VERSION : 0.1
   VAR_INPUT
      search_term : WString;
      search_array : Array[*] of WString[1];
   END_VAR
   VAR_TEMP
      _i : Int;
      _length_search_array : UDInt;
   END_VAR
BEGIN
   #_length_search_array := "Array.Any.Length"(#search_array);
   FOR #_i := 0 TO UDINT_TO_INT(#_length_search_array - 1) DO
       IF #search_term = #search_array[#_i] THEN
           #"Array.WString.Is_Element" := TRUE;
           RETURN;
       END_IF;
   END_FOR;
   #"Array.WString.Is_Element" := FALSE;
END_FUNCTION

FUNCTION "Array.Int.First_Occurance" : DInt   // FC220, SCL
{ S7_Optimized_Access := 'TRUE' }
VERSION : 0.1
   VAR_INPUT
      int_array : Array[*] of Int;
      search_term : Int;
   END_VAR
   VAR_TEMP
      _i : DInt;
      _length : UDInt;
   END_VAR
BEGIN
   REGION "NOTES"
       (* 
       This function returns the first occurance of the search term.
       This function meant for use with collapsed arrays.
       See "Array.Int.Collapse" for collapse functionality.
       *)
   END_REGION


   REGION "GET LENGTH OF INPUT ARRAY"
       #_length := "Array.Any.Length"(#int_array);
   END_REGION


   REGION "FIND FIRST SEARCH TERM, -1 IF NONE"
       (*
       Its worth noting that "Array.Int.Is_Element" could return the index of the search term
       as an output, saving the processor some work. 
       The rework is justified by increased encapsulation.
       The time complexity for "Array.Int.First_Occurance" remains O(n).
       *)
       IF NOT "Array.Int.Is_Element"(int_array := #int_array, search_term := #search_term) THEN
           #"Array.Int.First_Occurance" := -1;
           RETURN;
       END_IF;
       WHILE #int_array[#_i] <> #search_term AND DINT_TO_UDINT(#_i) < #_length DO
           #_i += 1;
       END_WHILE;
   END_REGION


   REGION _name_
       #"Array.Int.First_Occurance" := #_i;
   END_REGION
END_FUNCTION

FUNCTION "Array.WString.Fill" : Void   // FC243, SCL
{ S7_Optimized_Access := 'TRUE' }
VERSION : 0.1
   VAR_INPUT
      value : WString;
   END_VAR
   VAR_IN_OUT
      "array" : Array[*] of WString;
   END_VAR
   VAR_TEMP
      _length : Int;
      _i : Int;
   END_VAR
BEGIN
   #_length := UDINT_TO_INT("Array.Any.Length"(#array)) - 1;
   FOR #_i := 0 TO #_length DO
       #array[#_i] := #value;
   END_FOR;
   RETURN;
END_FUNCTION

FUNCTION "Array.WString.Search" : Int   // FC244, SCL
{ S7_Optimized_Access := 'TRUE' }
VERSION : 0.1
   VAR_INPUT
      "array" : Array[*] of WString;
      search_term : WString;
   END_VAR
   VAR_TEMP
      _i : Int;
      _length : Int;
   END_VAR
   // Ret_Val : index of search term. returns -1 if not found.
BEGIN
   REGION "SEARCH ARRAY"
       #_length := UDINT_TO_INT("Array.Any.Length"(#array)) - 1;
       FOR #_i := 0 TO #_length DO
           IF #array[#_i] <> #search_term THEN
               CONTINUE;
           END_IF;
           #"Array.WString.Search" := #_i;
           RETURN;
       END_FOR;
   END_REGION

   REGION "RETURN"
       #"Array.WString.Search" := "NULL_TOKEN";
       RETURN;
   END_REGION
END_FUNCTION

// folder: Utilities/Bool

FUNCTION "Bool.Animate" : USInt   // FC9, SCL
{ S7_Optimized_Access := 'TRUE' }
VERSION : 0.1
   VAR_INPUT
      true_color : USInt;
      false_color : USInt;
      evaluation_signal : Bool;
   END_VAR
   VAR_TEMP
      animate : USInt;
   END_VAR
BEGIN
   REGION "FALSE COLOR"
       IF NOT #evaluation_signal THEN
           #animate := #false_color;
       END_IF;
   END_REGION

   REGION "TRUE COLOR"
       IF #evaluation_signal THEN
           #animate := #true_color;
       END_IF;
   END_REGION

   REGION "FUNCTION RETURN"
       #"Bool.Animate" := #animate;
   END_REGION
END_FUNCTION

FUNCTION "Bool.Rising_Edge" : Bool   // FC177, SCL
{ S7_Optimized_Access := 'TRUE' }
VERSION : 0.1
   VAR_INPUT
      signal : Bool;
      old_signal : Bool;
   END_VAR
BEGIN
   #"Bool.Rising_Edge" := #signal AND NOT #old_signal;
END_FUNCTION

FUNCTION "Bool.Falling_Edge" : Bool   // FC178, SCL
{ S7_Optimized_Access := 'TRUE' }
VERSION : 0.1
   VAR_INPUT
      signal : Bool;
      old_signal : Bool;
   END_VAR
BEGIN
   #"Bool.Falling_Edge" := NOT #signal AND #old_signal;
END_FUNCTION

// folder: Utilities/DInt

FUNCTION "DInt.Clip.Maximum" : DInt   // FC224, SCL
{ S7_Optimized_Access := 'TRUE' }
VERSION : 0.1
   VAR_INPUT
      value : DInt;
      maximum : DInt;
   END_VAR
BEGIN
   IF #value > #maximum THEN
       #"DInt.Clip.Maximum" := #maximum;
       RETURN;
   END_IF;
   #"DInt.Clip.Maximum" := #value;
END_FUNCTION

FUNCTION "DInt.Clip.Minimum" : DInt   // FC225, SCL
{ S7_Optimized_Access := 'TRUE' }
VERSION : 0.1
   VAR_INPUT
      value : DInt;
      minimum : DInt;
   END_VAR
BEGIN
   IF #value < #minimum THEN
       #"DInt.Clip.Minimum" := #minimum;
       RETURN;
   END_IF;
   #"DInt.Clip.Minimum" := #value;
END_FUNCTION

FUNCTION "DInt.Clip.Range" : DInt   // FC227, SCL
{ S7_Optimized_Access := 'TRUE' }
VERSION : 0.1
   VAR_INPUT
      value : DInt;
      maximum : DInt;
      minimum : DInt;
   END_VAR
   VAR_TEMP
      _return : DInt;
   END_VAR
BEGIN
   #_return := #value;
   #_return := "DInt.Clip.Maximum"(value := #value, maximum := #minimum);
   #_return := "DInt.Clip.Minimum"(value := #value, minimum := #minimum);
   #"DInt.Clip.Range" := #_return;
END_FUNCTION

// folder: Utilities/Int

FUNCTION "Int.Value_Change" : Bool   // FC179, SCL
{ S7_Optimized_Access := 'TRUE' }
VERSION : 0.1
   VAR_INPUT
      value : Int;
      old_value : Int;
   END_VAR
BEGIN
   #"Int.Value_Change" := #value <> #old_value;
END_FUNCTION

FUNCTION "Int.Clip.Minimum" : Int   // FC222, SCL
{ S7_Optimized_Access := 'TRUE' }
VERSION : 0.1
   VAR_INPUT
      value : Int;
      minimum : Int;
   END_VAR
BEGIN
   IF #value < #minimum THEN
       #"Int.Clip.Minimum" := #minimum;
       RETURN;
   END_IF;
   #"Int.Clip.Minimum" := #value;
END_FUNCTION

FUNCTION "Int.Clip.Maximum" : Int   // FC223, SCL
{ S7_Optimized_Access := 'TRUE' }
VERSION : 0.1
   VAR_INPUT
      value : Int;
      maximum : Int;
   END_VAR
BEGIN
   IF #value > #maximum THEN
       #"Int.Clip.Maximum" := #maximum;
       RETURN;
   END_IF;
   #"Int.Clip.Maximum" := #value;
END_FUNCTION

FUNCTION "Int.Clip.Range" : Int   // FC226, SCL
{ S7_Optimized_Access := 'TRUE' }
VERSION : 0.1
   VAR_INPUT
      value : Int;
      maximum : Int;
      minimum : Int;
   END_VAR
   VAR_TEMP
      _return : Int;
   END_VAR
BEGIN
   #_return := #value;
   #_return := "Int.Clip.Maximum"(value := #_return, maximum := #maximum);
   #_return := "Int.Clip.Minimum"(value:=#_return, minimum:=#minimum);
   #"Int.Clip.Range" := #_return;
END_FUNCTION

// folder: Utilities/NavBar

FUNCTION_BLOCK "NavBar: Top"   // FB31, SCL
{ S7_Optimized_Access := 'TRUE' }
VERSION : 0.1
   VAR_INPUT
      hide : Bool;
      TABLE_LENGTH : DInt;
   END_VAR
   VAR_IN_OUT
      interface : "Push Button Data";
      first_row : DInt;
   END_VAR
   VAR
      "Get Button Feedback" : "Push Button: State Changes";
   END_VAR
   VAR_TEMP
      feedback : "Push Button Data: State Change Data";
   END_VAR
BEGIN
   REGION "PROCESS USER INPUT"
       #"Get Button Feedback"(interface := #interface,
                              state_changes := #feedback);
   END_REGION

   REGION "ANIMATIONS"

       REGION "COLOR"
           #interface.animate := "Bool.Animate"(true_color := "GREEN_LIGHT_BACKGROUND",
                                                false_color := "GRAY_BACKGROUND",
                                                evaluation_signal := #feedback.actuate.actual);
       END_REGION

       REGION "VISIBILITY"
           #interface.visible := NOT #hide;
       END_REGION

       REGION "ENABLED STATE"
           #interface.enable := NOT #hide;
       END_REGION

   END_REGION

   REGION "SET FIRST ROW"
       IF #feedback.actuate.rising THEN
           #first_row := 0;
       END_IF;
   END_REGION
END_FUNCTION_BLOCK

FUNCTION_BLOCK "NavBar: Bottom"   // FB32, SCL
{ S7_Optimized_Access := 'TRUE' }
VERSION : 0.1
   VAR_INPUT
      TABLE_LENGTH : DInt;
      VISIBLE_ROW_COUNT : DInt;
   END_VAR
   VAR_IN_OUT
      interface : "Push Button Data";
      first_row : DInt;
   END_VAR
   VAR
      "Get Button Feedback" : "Push Button: State Changes";
   END_VAR
   VAR_TEMP
      feedback : "Push Button Data: State Change Data";
   END_VAR
BEGIN
   REGION "PROCESS USER INPUT"
       #"Get Button Feedback"(interface := #interface,
                              state_changes := #feedback);
   END_REGION

   REGION "ANIMATIONS"

       REGION "COLOR"
           #interface.animate := "Bool.Animate"(true_color := "GREEN_LIGHT_BACKGROUND",
                                                false_color := "GRAY_BACKGROUND",
                                                evaluation_signal := #feedback.actuate.actual);
       END_REGION

       REGION "VISIBILITY"
           #interface.visible := TRUE;
       END_REGION

       REGION "ENABLED STATE"
           #interface.enable := TRUE;
       END_REGION

   END_REGION


   REGION "SET FIRST ROW"
       IF #feedback.actuate.rising THEN
           #first_row := #TABLE_LENGTH - #VISIBLE_ROW_COUNT;
       END_IF;
   END_REGION
END_FUNCTION_BLOCK

FUNCTION_BLOCK "NavBar: Page Up"   // FB36, SCL
{ S7_Optimized_Access := 'TRUE' }
VERSION : 0.1
   VAR_INPUT
      TABLE_LENGTH : DInt;
      VISIBLE_ROW_COUNT : DInt;
   END_VAR
   VAR_IN_OUT
      interface : "Push Button Data";
      first_row : DInt;
   END_VAR
   VAR
      "Get Button Feedback" : "Push Button: State Changes";
   END_VAR
   VAR_TEMP
      feedback : "Push Button Data: State Change Data";
   END_VAR
BEGIN
   REGION "PROCESS USER INPUT"
       #"Get Button Feedback"(interface := #interface,
                              state_changes := #feedback);
   END_REGION

   REGION "ANIMATIONS"

       REGION "COLOR"
           #interface.animate := "Bool.Animate"(true_color := "GREEN_LIGHT_BACKGROUND",
                                                false_color := "GRAY_BACKGROUND",
                                                evaluation_signal := #feedback.actuate.actual);
       END_REGION

       REGION "VISIBILITY"
           #interface.visible := TRUE;
       END_REGION

       REGION "ENABLED STATE"
           #interface.enable := TRUE;
       END_REGION

   END_REGION

   REGION "SET FIRST ROW"
       IF #feedback.actuate.rising THEN
           #first_row := "NavBar: Private: First Row"(first_row := #first_row,
                                                      offset := -1 * (#VISIBLE_ROW_COUNT + 1),
                                                      TABLE_LENGTH := #TABLE_LENGTH);
       END_IF;
   END_REGION
END_FUNCTION_BLOCK

FUNCTION_BLOCK "NavBar: Page Down"   // FB37, SCL
{ S7_Optimized_Access := 'TRUE' }
VERSION : 0.1
   VAR_INPUT
      TABLE_LENGTH : DInt;
      VISIBLE_ROW_COUNT : DInt;
   END_VAR
   VAR_IN_OUT
      interface : "Push Button Data";
      first_row : DInt;
   END_VAR
   VAR
      "Get Button Feedback" : "Push Button: State Changes";
   END_VAR
   VAR_TEMP
      feedback : "Push Button Data: State Change Data";
   END_VAR
BEGIN
   REGION "PROCESS USER INPUT"
       #"Get Button Feedback"(interface := #interface,
                              state_changes := #feedback);
   END_REGION

   REGION "ANIMATIONS"

       REGION "COLOR"
           #interface.animate := "Bool.Animate"(true_color := "GREEN_LIGHT_BACKGROUND",
                                                false_color := "GRAY_BACKGROUND",
                                                evaluation_signal := #feedback.actuate.actual);
       END_REGION

       REGION "VISIBILITY"
           #interface.visible := TRUE;
       END_REGION

       REGION "ENABLED STATE"
           #interface.enable := TRUE;
       END_REGION

   END_REGION

   REGION "SET FIRST ROW"
       IF #feedback.actuate.rising THEN
           #first_row := "NavBar: Private: First Row"(first_row := #first_row,
                                                      offset := #VISIBLE_ROW_COUNT + 1,
                                                      TABLE_LENGTH := #TABLE_LENGTH);
       END_IF;
   END_REGION
END_FUNCTION_BLOCK

FUNCTION_BLOCK "NavBar: Line Down"   // FB38, SCL
{ S7_Optimized_Access := 'TRUE' }
VERSION : 0.1
   VAR_INPUT
      TABLE_LENGTH : DInt;
   END_VAR
   VAR_IN_OUT
      interface : "Push Button Data";
      first_row : DInt;
   END_VAR
   VAR
      "Get Button Feedback" : "Push Button: State Changes";
   END_VAR
   VAR_TEMP
      feedback : "Push Button Data: State Change Data";
   END_VAR
BEGIN
   REGION "PROCESS USER INPUT"
       #"Get Button Feedback"(interface := #interface,
                              state_changes := #feedback);
   END_REGION

   REGION "ANIMATIONS"

       REGION "COLOR"
           #interface.animate := "Bool.Animate"(true_color := "GREEN_LIGHT_BACKGROUND",
                                                false_color := "GRAY_BACKGROUND",
                                                evaluation_signal := #feedback.actuate.actual);
       END_REGION

       REGION "VISIBILITY"
           #interface.visible := TRUE;
       END_REGION

       REGION "ENABLED STATE"
           #interface.enable := TRUE;
       END_REGION

   END_REGION

   REGION "SET FIRST ROW"
       IF #feedback.actuate.rising THEN
           #first_row := "NavBar: Private: First Row"(first_row := #first_row,
                                                      offset := 1,
                                                      TABLE_LENGTH := #TABLE_LENGTH);
       END_IF;
   END_REGION
END_FUNCTION_BLOCK

FUNCTION_BLOCK "NavBar: Line Up"   // FB39, SCL
{ S7_Optimized_Access := 'TRUE' }
VERSION : 0.1
   VAR_INPUT
      TABLE_LENGTH : DInt;
   END_VAR
   VAR_IN_OUT
      interface : "Push Button Data";
      first_row : DInt;
   END_VAR
   VAR
      "Get Button Feedback" : "Push Button: State Changes";
   END_VAR
   VAR_TEMP
      feedback : "Push Button Data: State Change Data";
   END_VAR
BEGIN
   REGION "PROCESS USER INPUT"
       #"Get Button Feedback"(interface := #interface,
                              state_changes := #feedback);
   END_REGION

   REGION "ANIMATIONS"

       REGION "COLOR"
           #interface.animate := "Bool.Animate"(true_color := "GREEN_LIGHT_BACKGROUND",
                                                false_color := "GRAY_BACKGROUND",
                                                evaluation_signal := #feedback.actuate.actual);
       END_REGION

       REGION "VISIBILITY"
           #interface.visible := TRUE;
       END_REGION

       REGION "ENABLED STATE"
           #interface.enable := TRUE;
       END_REGION

   END_REGION

   REGION "SET FIRST ROW"
       IF #feedback.actuate.rising THEN
           #first_row := "NavBar: Private: First Row"(first_row := #first_row,
                                                      offset := -1,
                                                      TABLE_LENGTH := #TABLE_LENGTH);
       END_IF;
   END_REGION
END_FUNCTION_BLOCK

FUNCTION_BLOCK "NavBar"   // FB40, SCL
{ S7_Optimized_Access := 'TRUE' }
VERSION : 0.1
   VAR_INPUT
      hide : Bool;
      TABLE_LENGTH : DInt := 49;
      VISIBLE_ROW_COUNT : DInt := 2;
   END_VAR
   VAR_IN_OUT
      interface : "Nav Bar Data";
      first_row : DInt;
   END_VAR
   VAR
      Top : "NavBar: Top";
      "Page Up" : "NavBar: Page Up";
      "Line Up" : "NavBar: Line Up";
      "Line Down" : "NavBar: Line Down";
      "Page Down" : "NavBar: Page Down";
      Bottom : "NavBar: Bottom";
   END_VAR
BEGIN
   REGION "BUFFER IN"
       "NavBar: Map HMI to PLC"(hmi := #interface.hmi,
                                plc := #interface.plc);
   END_REGION

   REGION "NAVBAR TOP "
       #Top(hide := #hide,
            TABLE_LENGTH := #TABLE_LENGTH,
            interface := #interface.plc.top,
            first_row := #first_row);
   END_REGION

   REGION "PAGE UP"
       #"Page Up"(TABLE_LENGTH := #TABLE_LENGTH,
                  VISIBLE_ROW_COUNT := #VISIBLE_ROW_COUNT,
                  interface := #interface.plc.pageUp,
                  first_row := #first_row);
   END_REGION

   REGION "LINE UP"
       #"Line Up"(TABLE_LENGTH := #TABLE_LENGTH,
                  interface := #interface.plc.lineUp,
                  first_row := #first_row);
   END_REGION

   REGION "LINE DOWN"
       #"Line Down"(TABLE_LENGTH := #TABLE_LENGTH,
                    interface := #interface.plc.lineDown,
                    first_row := #first_row);
   END_REGION

   REGION "PAGE DOWN"
       #"Page Down"(TABLE_LENGTH := #TABLE_LENGTH,
                    VISIBLE_ROW_COUNT := #VISIBLE_ROW_COUNT,
                    interface := #interface.plc.pageDown,
                    first_row := #first_row);
   END_REGION

   REGION "BOTTOM"
       #Bottom(TABLE_LENGTH := #TABLE_LENGTH,
               VISIBLE_ROW_COUNT := #VISIBLE_ROW_COUNT,
               interface := #interface.plc.bottom,
               first_row := #first_row);
   END_REGION

   REGION "BUFFER OUT"
       "NavBar: Map PLC to HMI"(plc := #interface.plc,
                                hmi := #interface.hmi);
   END_REGION
END_FUNCTION_BLOCK

FUNCTION "NavBar: Map HMI to PLC" : Void   // FC98, SCL
{ S7_Optimized_Access := 'TRUE' }
VERSION : 0.1
   VAR_INPUT
      hmi : "Nav Bar Data: HMI";
   END_VAR
   VAR_IN_OUT
      plc : "Nav Bar Data: PLC";
   END_VAR
BEGIN
   REGION "NOTES"
       // mapping is necessary because hmi faceplate data structures
       // cannot consist of embedded udts
   END_REGION


   REGION "TOP"
       #plc.top.actuate := #hmi.top_actuate;
       #plc.top.animate := #hmi.top_animate;
       #plc.top.enable := #hmi.top_enable;
       #plc.top.label := #hmi.top_label;
       #plc.top.listSelect := #hmi.top_list_select;
       #plc.top.visible := #hmi.top_visible;
   END_REGION


   REGION "PAGE UP"
       #plc.pageUp.actuate := #hmi.page_up_actuate;
       #plc.pageUp.animate := #hmi.page_up_animate;
       #plc.pageUp.enable := #hmi.page_up_enable;
       #plc.pageUp.label := #hmi.page_up_label;
       #plc.pageUp.listSelect := #hmi.page_up_list_select;
       #plc.pageUp.visible := #hmi.page_up_visible;
   END_REGION


   REGION "LINE UP"
       #plc.lineUp.actuate := #hmi.line_up_actuate;
       #plc.lineUp.animate := #hmi.line_up_animate;
       #plc.lineUp.enable := #hmi.line_up_enable;
       #plc.lineUp.label := #hmi.line_up_label;
       #plc.lineUp.listSelect := #hmi.line_up_list_select;
       #plc.lineUp.visible := #hmi.line_up_visible;
   END_REGION


   REGION "LINE DOWN"
       #plc.lineDown.actuate := #hmi.line_down_actuate;
       #plc.lineDown.animate := #hmi.line_down_animate;
       #plc.lineDown.enable := #hmi.line_down_enable;
       #plc.lineDown.label := #hmi.line_down_label;
       #plc.lineDown.listSelect := #hmi.line_down_list_select;
       #plc.lineDown.visible := #hmi.line_down_visible;
   END_REGION


   REGION "PAGE DOWN"
       #plc.pageDown.actuate := #hmi.page_down_actuate;
       #plc.pageDown.animate := #hmi.page_down_animate;
       #plc.pageDown.enable := #hmi.page_down_enable;
       #plc.pageDown.label := #hmi.page_down_label;
       #plc.pageDown.listSelect := #hmi.page_down_list_select;
       #plc.pageDown.visible := #hmi.page_down_visible;
   END_REGION


   REGION "BOTTOM"
       #plc.bottom.actuate := #hmi.bottom_actuate;
       #plc.bottom.animate := #hmi.bottom_animate;
       #plc.bottom.enable := #hmi.bottom_enable;
       #plc.bottom.label := #hmi.bottom_label;
       #plc.bottom.listSelect := #hmi.bottom_list_select;
       #plc.bottom.visible := #hmi.bottom_visible;
   END_REGION
END_FUNCTION

FUNCTION "NavBar: Map PLC to HMI" : Void   // FC99, SCL
{ S7_Optimized_Access := 'TRUE' }
VERSION : 0.1
   VAR_INPUT
      plc : "Nav Bar Data: PLC";
   END_VAR
   VAR_IN_OUT
      hmi : "Nav Bar Data: HMI";
   END_VAR
BEGIN
   REGION "NOTES"
       // mapping is necessary because hmi faceplate data structures
       // cannot consist of embedded udts
   END_REGION


   REGION "TOP"
       //#hmi.top_actuate := #plc.top.actuate;
       #hmi.top_animate := #plc.top.animate;
       #hmi.top_enable := #plc.top.enable;
       #hmi.top_label := #plc.top.label;
       #hmi.top_list_select := #plc.top.listSelect;
       #hmi.top_visible := #plc.top.visible;
   END_REGION


   REGION "PAGE UP"
       //#hmi.page_up_actuate := #plc.pageUp.actuate;
       #hmi.page_up_animate := #plc.pageUp.animate;
       #hmi.page_up_enable := #plc.pageUp.enable;
       #hmi.page_up_label := #plc.pageUp.label;
       #hmi.page_up_list_select := #plc.pageUp.listSelect;
       #hmi.page_up_visible := #plc.pageUp.visible;
   END_REGION


   REGION "LINE UP"
       //#hmi.line_up_actuate := #plc.lineUp.actuate;
       #hmi.line_up_animate := #plc.lineUp.animate;
       #hmi.line_up_enable := #plc.lineUp.enable;
       #hmi.line_up_label := #plc.lineUp.label;
       #hmi.line_up_list_select := #plc.lineUp.listSelect;
       #hmi.line_up_visible := #plc.lineUp.visible;
   END_REGION


   REGION "LINE DOWN"
       //#hmi.line_down_actuate := #plc.lineDown.actuate;
       #hmi.line_down_animate := #plc.lineDown.animate;
       #hmi.line_down_enable := #plc.lineDown.enable;
       #hmi.line_down_label := #plc.lineDown.label;
       #hmi.line_down_list_select := #plc.lineDown.listSelect;
       #hmi.line_down_visible := #plc.lineDown.visible;
   END_REGION


   REGION "PAGE DOWN"
       //#hmi.page_down_actuate := #plc.pageDown.actuate;
       #hmi.page_down_animate := #plc.pageDown.animate;
       #hmi.page_down_enable := #plc.pageDown.enable;
       #hmi.page_down_label := #plc.pageDown.label;
       #hmi.page_down_list_select := #plc.pageDown.listSelect;
       #hmi.page_down_visible := #plc.pageDown.visible;
   END_REGION

   REGION "BOTTOM"
       //#hmi.bottom_actuate := #plc.bottom.actuate;
       #hmi.bottom_animate := #plc.bottom.animate;
       #hmi.bottom_enable := #plc.bottom.enable;
       #hmi.bottom_label := #plc.bottom.label;
       #hmi.bottom_list_select := #plc.bottom.listSelect;
       #hmi.bottom_visible := #plc.bottom.visible;
   END_REGION
END_FUNCTION

FUNCTION "NavBar: Private: First Row" : DInt   // FC180, SCL
{ S7_Optimized_Access := 'TRUE' }
VERSION : 0.1
   VAR_INPUT
      first_row : DInt;
      offset : DInt;
      TABLE_LENGTH : DInt;
   END_VAR
   VAR_TEMP
      ret : DInt;
   END_VAR
BEGIN
   REGION "DESCRIPTION"
       (*
       The new first row of the table is calculated from the offset. 
       Rollover and rollunder are resolved for the first row.
       *)
   END_REGION

   REGION "COPY TO INTERNAL"
       #ret := #first_row + #offset;
   END_REGION

   REGION "ROLLUNDER"
       IF #ret < 0 THEN
           #ret := #ret + #TABLE_LENGTH + 1;
       END_IF;
   END_REGION

   REGION "ROLLOVER"
       IF #ret > #TABLE_LENGTH THEN
           #ret := #ret - #TABLE_LENGTH - 1;
       END_IF;
   END_REGION

   REGION "OUTPUT"
       #"NavBar: Private: First Row" := #ret;
   END_REGION
END_FUNCTION

// folder: Utilities/Part Number

FUNCTION "Part_Number.Parse_Code" : Void   // FC34, SCL
{ S7_Optimized_Access := 'TRUE' }
VERSION : 0.1
   VAR_INPUT
      code : DInt;
   END_VAR
   VAR_OUTPUT
      code_left : DInt;
      code_right : DInt;
   END_VAR
BEGIN
   IF #code > 0 THEN
       #code_left := #code / 1000;
       #code_right := #code - #code / 1000 * 1000;
   ELSE
       #code_left := 0;
       #code_right := 0;
   END_IF;
END_FUNCTION

FUNCTION "Part_Number.Code_to_WString" : WString   // FC37, SCL
{ S7_Optimized_Access := 'TRUE' }
VERSION : 0.1
   VAR_INPUT
      pnLib : "Recipe: PN Text Library";
      pnCode : DInt;
   END_VAR
   VAR_TEMP
      pnLeft : DInt;
      pnRight : DInt;
      output : WString;
   END_VAR
   VAR CONSTANT
      newLine : WString := WSTRING#'$L';
   END_VAR
BEGIN
   REGION "PARSE CODE"
       "Part_Number.Parse_Code"(code := #pnCode,
                                 code_left => #pnLeft,
                                 code_right => #pnRight);
   END_REGION

   REGION "SINGLE LINE PN"
       IF "Part_Number.Is_Single"(#pnCode) THEN
           #output := #pnLib.pnText[#pnLeft];
       END_IF;
   END_REGION

   REGION "DOUBLE LINE PN"
       IF "Part_Number.Is_Double"(#pnCode) THEN
           #output := CONCAT_WSTRING(IN1 := #pnLib.pnText[#pnLeft],
                                     IN2 := #newLine,
                                     IN3 := #pnLib.pnText[#pnRight]);
       END_IF;
   END_REGION

   REGION "OUTPUT"
       #"Part_Number.Code_to_WString" := #output;
   END_REGION
END_FUNCTION

FUNCTION "Part_Number.Is_Double" : Bool   // FC153, SCL
{ S7_Optimized_Access := 'TRUE' }
VERSION : 0.1
   VAR_INPUT
      code : DInt;
   END_VAR
   VAR_TEMP
      code_left : DInt;
      code_right : DInt;
      ret : Bool;
   END_VAR
BEGIN
   REGION "NOTES"
       (*
       Double codes have a non-zero right hand component.
       Structure: XXXYYY
       XXX: left code, used for single and double codes
       YYY: right code, only used for double codes
       Last Edit: 2021-10-07
       *)
   END_REGION

   REGION "PROCESS CODE"
       "Part_Number.Parse_Code"(code := #code,
                                code_left => #code_left,
                                code_right => #code_right);
   END_REGION

   REGION "CHECK FOR DOUBLE CODE"
       IF #code_right > 0 THEN
           #ret := TRUE;
       END_IF;
   END_REGION

   REGION "RETURN" 
       #"Part_Number.Is_Double" := #ret;
   END_REGION
END_FUNCTION

FUNCTION "Part_Number.Is_Single" : Bool   // FC154, SCL
{ S7_Optimized_Access := 'TRUE' }
VERSION : 0.1
   VAR_INPUT
      code : DInt;
   END_VAR
   VAR_TEMP
      code_left : DInt;
      code_right : DInt;
      ret : Bool;
   END_VAR
BEGIN
   REGION "NOTES"
       (*
       Double codes have a non-zero right hand component.
       Structure:
       XXXYYY
       XXX: left code, used for single and double codes
       YYY: right code, only used for double codes
       Last Edit: 2021-10-07
       *)
   END_REGION

   REGION "PROCESS CODE"
       "Part_Number.Parse_Code"(code := #code,
                                code_left => #code_left,
                                code_right => #code_right);
   END_REGION

   REGION "CHECK FOR DOUBLE CODE"
       IF #code_right = 0 THEN
           #ret := TRUE;
       END_IF;
   END_REGION

   REGION "RETURN" 
       #"Part_Number.Is_Single" := #ret;
   END_REGION
END_FUNCTION

FUNCTION "Part_Number.WString_to_Code" : DInt   // FC240, SCL
{ S7_Optimized_Access := 'TRUE' }
VERSION : 0.1
   VAR_INPUT
      part_number : WString;
   END_VAR
   VAR_IN_OUT
      pn_library : "Recipe: PN Text Library";
   END_VAR
   VAR_TEMP
      _in_library : Bool;
      _library_full : Bool;
      _part_numbers : Array[0..1] of WString;
      _partial_pn_code : DInt;
      _pn_count : Int;
      _pn_code : DInt;
   END_VAR
   VAR CONSTANT
      OUT_OF_MEMORY : DInt := 999;
   END_VAR
BEGIN
   REGION "DATA PREP""
       "Part_Number.Split_PNs"(part_number := #part_number,
                               part_numbers := #_part_numbers);
       #_pn_count := "Part_Number.Count_PNs"(#_part_numbers);
   END_REGION


   REGION "NO PART NUMBERS ENTERED"
       IF #_pn_count = 0 THEN
           #"Part_Number.WString_to_Code" := 0;
           RETURN;
       END_IF;
   END_REGION


   REGION "CHECK FIRST PN CODE"
       #_pn_code := "Part_Number_Library.Search"(pn_library := #pn_library,
                                                 search_term := #_part_numbers[0]);
       #_in_library := "Part_Number.In_Library"(#_pn_code);
       #_library_full := "Part_Number_Library.Is_Full"(#pn_library);
   END_REGION


   REGION "FIRST PN CODE IN LIBRARY"
       IF #_in_library THEN
           #_pn_code *= 1_000;
       END_IF;
   END_REGION


   REGION "FIRST PN NOT IN LIBRARY, NO SPACE"
       IF NOT #_in_library AND #_library_full THEN
           #_pn_code := #OUT_OF_MEMORY * 1_000;
       END_IF;
   END_REGION


   REGION "FIRST PN NOT IN LIBRARY, SPACE"
       IF NOT #_in_library AND NOT #_library_full THEN
           #_pn_code := 1_000 * "Part_Number_Library.Add_PN"(pn := #_part_numbers[0],
                                                             pn_library := #pn_library);
       END_IF;
   END_REGION


   REGION "RETURN SINGLE PN CODE"
       IF #_pn_count = 1 THEN
           #"Part_Number.WString_to_Code" := #_pn_code;
           RETURN;
       END_IF;
   END_REGION


   REGION "CHECK SECOND PN CODE"
       #_partial_pn_code := "Part_Number_Library.Search"(pn_library := #pn_library,
                                                         search_term := #_part_numbers[1]);
       #_in_library := "Part_Number.In_Library"(#_partial_pn_code);
       #_library_full := "Part_Number_Library.Is_Full"(#pn_library);
   END_REGION


   REGION "SECOND PN CODE IN LIBRARY"
       IF #_in_library THEN
           #"Part_Number.WString_to_Code" := #_pn_code + #_partial_pn_code;
           RETURN;
       END_IF;
   END_REGION


   REGION "FIRST PN NOT IN LIBRARY, NO SPACE"
       IF NOT #_in_library AND #_library_full THEN
           #"Part_Number.WString_to_Code" := #_pn_code + #OUT_OF_MEMORY;
           RETURN;
       END_IF;
   END_REGION


   REGION "FIRST PN NOT IN LIBRARY, SPACE"
       IF NOT #_in_library AND NOT #_library_full THEN
           #_pn_code += "Part_Number_Library.Add_PN"(pn := #_part_numbers[0],
                                                     pn_library := #pn_library);
           #"Part_Number.WString_to_Code" := #_pn_code;
           RETURN;
       END_IF;
   END_REGION


   #"Part_Number.WString_to_Code" := 0;
   RETURN;
END_FUNCTION

FUNCTION "Part_Number.Count_PNs" : Int   // FC252, SCL
{ S7_Optimized_Access := 'TRUE' }
VERSION : 0.1
   VAR_INPUT
      part_numbers : Array[0..1] of WString;
   END_VAR
   VAR CONSTANT
      NULL : WString := WSTRING#'//';
      BLANK : WString := WSTRING#'';
   END_VAR
BEGIN
   IF #part_numbers[0] = #NULL THEN
       #"Part_Number.Count_PNs" := 0;
       RETURN;
   END_IF;

   IF #part_numbers[0] = #BLANK THEN
       #"Part_Number.Count_PNs" := 0;
       RETURN;
   END_IF;

   IF #part_numbers[1] = #NULL THEN
       #"Part_Number.Count_PNs" := 1;
       RETURN;
   END_IF;

   IF #part_numbers[1] = #BLANK THEN
       #"Part_Number.Count_PNs" := 1;
       RETURN;
   END_IF;

   #"Part_Number.Count_PNs" := 2;
   RETURN;
END_FUNCTION

FUNCTION "Part_Number.In_Library" : Bool   // FC253, SCL
{ S7_Optimized_Access := 'TRUE' }
VERSION : 0.1
   VAR_INPUT
      pn_code : DInt;
   END_VAR
BEGIN
   IF #pn_code = "NULL_TOKEN" THEN
       #"Part_Number.In_Library" := FALSE;
       RETURN;
   END_IF;
   #"Part_Number.In_Library" := TRUE;
   RETURN;
END_FUNCTION

FUNCTION "Part_Number.Split_PNs" : Void   // FC254, SCL
{ S7_Optimized_Access := 'TRUE' }
VERSION : 0.1
   VAR_INPUT
      part_number : WString;
   END_VAR
   VAR_IN_OUT
      part_numbers : Array[0..1] of WString;
   END_VAR
   VAR_TEMP
      _part_numbers : Array[0..1] of WString;
   END_VAR
   VAR CONSTANT
      NEW_LINE : WString := WSTRING#'$L';
      NULL : WString := WSTRING#'//';
   END_VAR
BEGIN
   "Array.WString.Fill"(value := #NULL,
                        array := #_part_numbers);
   "WString.Split_Single"(wstring_in := #part_number,
                          delimeter := #NEW_LINE,
                          "pointer" := 0,
                          sub_strings := #_part_numbers);
   #part_numbers := #_part_numbers;
END_FUNCTION

// folder: Utilities/Part Number Library

FUNCTION "Part_Number_Library.Is_Full" : Bool   // FC250, SCL
{ S7_Optimized_Access := 'TRUE' }
VERSION : 0.1
   VAR_INPUT
      pn_library : "Recipe: PN Text Library";
   END_VAR
   VAR_TEMP
      _first_null : DInt;
   END_VAR
   VAR CONSTANT
      NULL_STRING : WString := WSTRING#'//';
   END_VAR
BEGIN
   #_first_null := "Part_Number_Library.Search"(pn_library := #pn_library,
                                                search_term := #NULL_STRING);
   IF #_first_null = "NULL_TOKEN" THEN
       #"Part_Number_Library.Is_Full" := TRUE;
       RETURN;
   END_IF;

   #"Part_Number_Library.Is_Full" := FALSE;
   RETURN;
END_FUNCTION

FUNCTION "Part_Number_Library.Add_PN" : DInt   // FC251, SCL
{ S7_Optimized_Access := 'TRUE' }
VERSION : 0.1
   VAR_INPUT
      pn : WString;
   END_VAR
   VAR_IN_OUT
      pn_library : "Recipe: PN Text Library";
   END_VAR
   VAR_TEMP
      _index : DInt;
   END_VAR
   VAR CONSTANT
      NULL_STRING : WString := WSTRING#'//';
   END_VAR
BEGIN
   #_index := "Part_Number_Library.Search"(pn_library := #pn_library,
                                           search_term := #NULL_STRING);
   #pn_library.pnText[#_index] := #pn;
   #"Part_Number_Library.Add_PN" := #_index;
END_FUNCTION

FUNCTION "Part_Number_Library.Search" : Int   // FC255, SCL
{ S7_Optimized_Access := 'TRUE' }
VERSION : 0.1
   VAR_INPUT
      pn_library : "Recipe: PN Text Library";
      search_term : WString;
   END_VAR
   VAR_TEMP
      _array : Array[0..#MAX_ELEMENTS] of WString;
      _slices : Int;
      _slice : Int;
      _internal_length : Int;
      _external_length : Int;
      _search_result : Int;
   END_VAR
   VAR CONSTANT
      MAX_ELEMENTS : Int := 24;
   END_VAR
BEGIN
   REGION "NOTES"
       (*
           Why is this necessary?
               Unfortunately, dynamically sized arrays of wstring data type cannot accept
               wstrings of a declared length (e.x. the input parameter array[*] of 
               wstring[10] cannot exist). We need this wrapper function so that we can 
               copy wstrings of a declared length to an array of wstrings of default 
               length. Once copied, this array can be passed into the wstring search 
               function. However, there is only 16k of local memory to store the array of
               wstrings of default length. The pn text library can store up to 1000 part 
               numbers. If we were to copy all 1000, we would need 500k of memory. So, we 
               must slice the pn library into chunks and search them.
           Why are part number text wstrings a declared length?
               The declared lenght was necessary to fit a reasonable number of part 
               numbers into retentive memory.
       *)
   END_REGION


   REGION "SETUP"
       #_internal_length := UDINT_TO_INT("Array.Any.Length"(#_array));
       #_external_length := UDINT_TO_INT("Array.Any.Length"(#pn_library.pnText));
       #_slices := #_external_length / #_internal_length - 1;
   END_REGION


   REGION "REPEAT FOR EACH SLICE OF EXTERNAL ARRAY"
       FOR #_slice := 0 TO #_slices DO
           "Part_Number_Library.Search.Map_to_Internal_Array"(pn_library := #pn_library,
                                                              slice_number := #_slice,
                                                              internal_array := #_array);
           #_search_result := "Array.WString.Search"(array := #_array,
                                                     search_term := #search_term);
           IF #_search_result <> "NULL_TOKEN" THEN
               #"Part_Number_Library.Search" := #_search_result + #_slice * #_internal_length;
               RETURN;
           END_IF;
       END_FOR;
   END_REGION

   REGION "RETURN"
       #"Part_Number_Library.Search" := "NULL_TOKEN";
       RETURN;
   END_REGION
END_FUNCTION

FUNCTION "Part_Number_Library.Search.Map_to_Internal_Array" : Void   // FC256, SCL
{ S7_Optimized_Access := 'TRUE' }
VERSION : 0.1
   VAR_INPUT
      pn_library : "Recipe: PN Text Library";
      slice_number : Int;
   END_VAR
   VAR_IN_OUT
      internal_array : Array[*] of WString;
   END_VAR
   VAR_TEMP
      _i : Int;
      _length : Int;
      _p : Int;
   END_VAR
BEGIN
   #_length := UDINT_TO_INT("Array.Any.Length"(#internal_array));
   FOR #_i := 0 TO #_length - 1 DO
       #_p := #_i + #slice_number * #_length;
       #internal_array[#_i] := #pn_library.pnText[#_p];
   END_FOR;
END_FUNCTION

// folder: Utilities/Screen Objects

FUNCTION "Cell_Data.Hide" : "Cell Data"   // FC209, SCL
{ S7_Optimized_Access := 'TRUE' }
VERSION : 0.1
BEGIN
   #"Cell_Data.Hide".animate := "INVISIBLE";
   #"Cell_Data.Hide".data := "BLANK";
   #"Cell_Data.Hide".visibility := "HIDE";
END_FUNCTION

FUNCTION "Cell_Data.Show" : "Cell Data"   // FC216, SCL
{ S7_Optimized_Access := 'TRUE' }
VERSION : 0.1
   VAR_INPUT
      animate : Int;
      data : WString;
   END_VAR
   VAR_TEMP
      _ret : "Cell Data";
   END_VAR
BEGIN
   #_ret.animate := #animate;
   #_ret.data := #data;
   #_ret.visibility := "SHOW";
   #"Cell_Data.Show" := #_ret;
END_FUNCTION

// folder: Utilities/Selected Buttons

FUNCTION "Selected_Buttons.Indices" : Void   // FC246, SCL
{ S7_Optimized_Access := 'TRUE' }
VERSION : 0.1
   VAR_INPUT
      selected_buttons : "Selected Buttons";
   END_VAR
   VAR_IN_OUT
      selected_stations_indices : Array[*] of Int;
   END_VAR
   VAR_TEMP
      _i : Int;
      _length : Int;
      _resized_bool_array : Array[0..999] of Bool;
   END_VAR
BEGIN
   #_length := UDINT_TO_INT("Array.Any.Length"(#selected_buttons.btns)) - 1;
   FOR #_i := 0 TO #_length DO
       #_resized_bool_array[#_i] := #selected_buttons.btns[#_i];
   END_FOR;
   "Array.Bool.True_Indices"(array_of_bool := #_resized_bool_array,
                             list_of_indices := #selected_stations_indices);

   #selected_stations_indices[0] := #selected_stations_indices[0];
   #selected_stations_indices[1] := #selected_stations_indices[1];
   #selected_stations_indices[2] := #selected_stations_indices[2];
   #selected_stations_indices[3] := #selected_stations_indices[3];
   #selected_stations_indices[4] := #selected_stations_indices[4];
   #selected_stations_indices[5] := #selected_stations_indices[5];
   #selected_stations_indices[6] := #selected_stations_indices[6];
   #selected_stations_indices[7] := #selected_stations_indices[7];


   FOR #_i := 0 TO #_length DO
       IF #selected_stations_indices[#_i] = "NULL_TOKEN" THEN
           CONTINUE;
       END_IF;
       #selected_stations_indices[#_i] := "KP8.DURL_to_LRUD"(#selected_stations_indices[#_i]);
   END_FOR;

   #selected_stations_indices[0] := #selected_stations_indices[0];
   #selected_stations_indices[1] := #selected_stations_indices[1];
   #selected_stations_indices[2] := #selected_stations_indices[2];
   #selected_stations_indices[3] := #selected_stations_indices[3];
   #selected_stations_indices[4] := #selected_stations_indices[4];
   #selected_stations_indices[5] := #selected_stations_indices[5];
   #selected_stations_indices[6] := #selected_stations_indices[6];
   #selected_stations_indices[7] := #selected_stations_indices[7];
END_FUNCTION

// folder: Utilities/Selected Stations

FUNCTION "Selected_Stations.Indices" : Void   // FC245, SCL
{ S7_Optimized_Access := 'TRUE' }
VERSION : 0.1
   VAR_INPUT
      selected_stations : "Selected Stations";
   END_VAR
   VAR_IN_OUT
      selected_stations_indices : Array[*] of Int;
   END_VAR
   VAR_TEMP
      _i : Int;
      _length : Int;
      _resized_array : Array[0..999] of Bool;
   END_VAR
BEGIN
   FOR #_i := 0 TO "STATION_COUNT" DO
       #_resized_array[#_i] := #selected_stations.stns[#_i];
   END_FOR;
   "Array.Bool.True_Indices"(array_of_bool := #_resized_array,
                             list_of_indices := #selected_stations_indices);
END_FUNCTION

// folder: Utilities/String

FUNCTION "Strip Sign" : WString   // FC3, SCL
{ S7_Optimized_Access := 'TRUE' }
VERSION : 0.1
   VAR_INPUT
      WString : WString;
   END_VAR
   VAR_TEMP
      Length : Int;
      "String Box" : WString;
      "Test Character" : WString;
   END_VAR
   VAR CONSTANT
      "+" : WChar := WCHAR#'+';
      "-" : WChar := WCHAR#'-';
   END_VAR
BEGIN
   #"String Box" := #WString;
   #"Test Character" := LEFT_WSTRING(IN := #"String Box",
                                     L := 1);
   IF #"Test Character" = #"+" OR #"Test Character" = #"-" THEN
       #Length := LEN(#"String Box");
       #"String Box" := RIGHT_WSTRING(IN := #"String Box", L := #Length - 1);

   END_IF;
   #"Strip Sign" := #"String Box";
END_FUNCTION

FUNCTION "Add Leading" : WString   // FC4, SCL
{ S7_Optimized_Access := 'TRUE' }
VERSION : 0.1
   VAR_INPUT
      "Leading Character" : WChar;
      "Desired Length" : USInt;
      "String" : WString;
   END_VAR
   VAR_TEMP
      Length : Int;
      "String Box" : WString;
   END_VAR
BEGIN
   #"String Box" := #String;
   #Length := LEN(#"String Box");

   WHILE #Length < #"Desired Length" DO
       #"String Box" := CONCAT_WSTRING(IN1 := #"Leading Character",
                                       IN2 := #"String Box");
       #Length := LEN(#"String Box");
   END_WHILE;

   #"Add Leading" := #"String Box";
END_FUNCTION

FUNCTION "WString.Word_Wrap_Depricated" : WString   // FC28, SCL
{ S7_Optimized_Access := 'TRUE' }
VERSION : 0.1
   VAR_INPUT
      stringIn : WString;
      maxLength : Int;
   END_VAR
   VAR_TEMP
      length : Int;
      lineBox : Array[0..#limitLines] of WString["LONG_STRING_LENGTH"];
      ret : WString;
      stringBox : Array[0..#limitString] of WString["LONG_STRING_LENGTH"];
   END_VAR
   VAR CONSTANT
      space : WString := WSTRING#' ';
      blank : WString;
      lineBreak : WString := WSTRING#'$L';
      limitString : Int := 49;
      limitLines : Int := 9;
   END_VAR
BEGIN
   REGION "GET LENGTH"
       #length := LEN(#stringIn);
   END_REGION

   REGION "NO WRAP NECESSARY"
       IF #length <= #maxLength THEN
           #ret := #stringIn;
       END_IF;
   END_REGION


   REGION "EXECUTE WORD WRAP"
       IF #length > #maxLength THEN

           "Explode"(stringIn := #stringIn,
                     explodedString := #stringBox);

           "WString.Word_Wrap_Depricated.Construct_Line"(stringBox := #stringBox,
                                       lineBox := #lineBox,
                                       maxLength := #maxLength);

           #ret := "WString.Word_Wrap_Depricated.Concat_Lines"(#lineBox);

       END_IF;
   END_REGION

   REGION "RETURN"
       #"WString.Word_Wrap_Depricated" := #ret;
   END_REGION
END_FUNCTION

FUNCTION "Trim" : WString   // FC29, SCL
{ S7_Optimized_Access := 'TRUE' }
VERSION : 0.1
   VAR_INPUT
      wString : WString;
   END_VAR
   VAR_TEMP
      ret : WString;
   END_VAR
   VAR CONSTANT
      space : WString := WSTRING#' ';
   END_VAR
BEGIN
   #ret := #wString;
   WHILE LEFT(IN := #ret, L := 1) = #space DO
       #ret := RIGHT(IN := #ret, L := LEN(#ret) - 1);
   END_WHILE;
   WHILE RIGHT(IN := #ret, L := 1) = #space DO
       #ret := LEFT(IN := #ret, L := LEN(#ret) - 1);
   END_WHILE;
   #Trim := #ret;
END_FUNCTION

FUNCTION "Upper" : Void   // FC49, SCL
{ S7_Optimized_Access := 'TRUE' }
VERSION : 0.1
   VAR_IN_OUT
      "string" : Variant;
   END_VAR
   VAR_TEMP
      "type" : Bool;
      stringBox : String;
      status : Int;
      wStringBox : WString;
      charArr : Array[0..255] of Char;
      cntChar : UInt;
      pChar : Int;
   END_VAR
   VAR CONSTANT
      asciiLow : Char := 'a';
      asciiHigh : Char := 'z';
      asciiCaseOffset : Int := 32;
   END_VAR
BEGIN
   IF TypeOf(#string) = String THEN
       #status := MOVE_BLK_VARIANT(SRC := #string,
                                   COUNT := 1,
                                   SRC_INDEX := 0,
                                   DEST_INDEX := 0,
                                   DEST => #stringBox);
   ELSIF TypeOf(#string) = WString THEN
       #status := MOVE_BLK_VARIANT(SRC := #string,
                                   COUNT := 1,
                                   SRC_INDEX := 0,
                                   DEST_INDEX := 0,
                                   DEST => #wStringBox);
       #stringBox := WSTRING_TO_STRING(#wStringBox);
   ELSE
       RETURN;
   END_IF;

   Strg_TO_Chars(Strg := #stringBox,
                 pChars := 0,
                 Cnt => #cntChar,
                 Chars := #charArr);

   FOR #pChar := 0 TO UINT_TO_INT(#cntChar) - 1 DO
       IF #asciiLow <= #charArr[#pChar] AND #charArr[#pChar] <= #asciiHigh THEN
           #charArr[#pChar] := INT_TO_CHAR(CHAR_TO_INT(#charArr[#pChar]) - #asciiCaseOffset);
       END_IF;
   END_FOR;

   Chars_TO_Strg(Chars := #charArr,
                 pChars := 0,
                 Cnt := #cntChar,
                 Strg => #stringBox);

   IF TypeOf(#string) = String THEN
       #status := MOVE_BLK_VARIANT(SRC := #stringBox,
                                   COUNT := 1,
                                   SRC_INDEX := 0,
                                   DEST_INDEX := 0,
                                   DEST => #string);
   ELSIF TypeOf(#string) = WString THEN
       #wStringBox := STRING_TO_WSTRING(#stringBox);
       #status := MOVE_BLK_VARIANT(SRC := #wStringBox,
                                   COUNT := 1,
                                   SRC_INDEX := 0,
                                   DEST_INDEX := 0,
                                   DEST => #string);
   END_IF;
END_FUNCTION

FUNCTION "Explode" : Void   // FC73, SCL
{ S7_Optimized_Access := 'TRUE' }
VERSION : 0.1
   VAR_INPUT
      stringIn : WString;
   END_VAR
   VAR_IN_OUT
      explodedString : Variant;
   END_VAR
   VAR_TEMP
      charBox : Array[0..#lmtChar] of WChar;
      count : DInt;
      pChar : Int;
      pStringBox : Int;
      stringBox : Array[0..#lmtString] of WString["LONG_STRING_LENGTH"];
      status : DInt;
   END_VAR
   VAR CONSTANT
      space : WString := WSTRING#' ';
      blank : WString;
      lineBreak : WString := WSTRING#'$L';
      lmtString : Int := 49;
      lmtChar : Int := 999;
   END_VAR
BEGIN
   Strg_TO_Chars(Strg := #stringIn,
                 pChars := 0,
                 Cnt => #count,
                 Chars := #charBox);

   FOR #pChar := 0 TO #count DO

       IF #charBox[#pChar] = #space THEN
           IF #charBox[#pChar + 1] = #space THEN
               EXIT;
           END_IF;
       END_IF;

       IF #pChar = 0 THEN
           #stringBox[#pStringBox] := #charBox[#pChar];
       END_IF;

       IF #pChar >= 1 THEN
           #stringBox[#pStringBox] := CONCAT_WSTRING(IN1 := #stringBox[#pStringBox],
                                                     IN2 := #charBox[#pChar]);
       END_IF;

       IF #charBox[#pChar] = #space THEN
           #stringBox[#pStringBox] := "Trim"(#stringBox[#pStringBox]);
           #pStringBox := #pStringBox + 1;
       END_IF;

       IF #charBox[#pChar] = #lineBreak THEN
           #stringBox[#pStringBox] := LEFT(IN := #stringBox[#pStringBox],
                                           L := LEN(#stringBox[#pStringBox]) - 1);
           #pStringBox := #pStringBox + 1;
           #stringBox[#pStringBox] := #lineBreak;
           #pStringBox := #pStringBox + 1;
       END_IF;

   END_FOR;

   #status := MOVE_BLK_VARIANT(SRC := #stringBox,
                               COUNT := INT_TO_UDINT(#pStringBox)+1,
                               SRC_INDEX :=0,
                               DEST_INDEX := 0,
                               DEST => #explodedString);
END_FUNCTION

FUNCTION "WString.Word_Wrap_Depricated.Construct_Line" : Void   // FC74, SCL
{ S7_Optimized_Access := 'TRUE' }
VERSION : 0.1
   VAR_INPUT
      stringBox : Array[0..#limitString] of WString["LONG_STRING_LENGTH"];
      maxLength : Int;
   END_VAR
   VAR_IN_OUT
      lineBox : Array[0..#limitLines] of WString["LONG_STRING_LENGTH"];
   END_VAR
   VAR_TEMP
      _lineBox : Array[0..#limitLines] of WString["LONG_STRING_LENGTH"];
      pString : Int;
      pLineBox : Int;
      lengthTest : WString;
   END_VAR
   VAR CONSTANT
      space : WString := WSTRING#' ';
      blank : WString;
      lineBreak : WString := WSTRING#'$L';
      limitString : Int := 49;
      limitLines : Int := 9;
   END_VAR
BEGIN
   REGION "FOR EACH STRING IN STRING LIST"
       FOR #pString := 0 TO #limitString DO

           REGION "END OF STRING LIST"
               IF #stringBox[#pString] = #blank THEN
                   IF #stringBox[#pString + 1] = #blank THEN
                       #_lineBox[#pLineBox] := "Trim"(#_lineBox[#pLineBox]);
                       #lineBox := #_lineBox;
                       RETURN;
                   END_IF;
               END_IF;
           END_REGION

           REGION "ON NEW LINE CHARACTER"
               IF #stringBox[#pString] = #lineBreak THEN
                   #_lineBox[#pLineBox] := "Trim"(#_lineBox[#pLineBox]);
                   #pLineBox := #pLineBox + 1;
                   #_lineBox[#pLineBox] := #lineBreak;
                   #pLineBox := #pLineBox + 1;
               END_IF;
           END_REGION

           REGION "BUILD EACH LINE"
               IF #stringBox[#pString] <> #lineBreak THEN

                   REGION "FIRST ELEMENT EDGE CASE"
                       IF #pString = 0 THEN
                           #lengthTest := #stringBox[#pString];
                       END_IF;
                   END_REGION

                   REGION "BUILT TEST STRING"
                       IF #pString >= 1 THEN
                           #lengthTest := CONCAT_WSTRING(IN1 := #_lineBox[#pLineBox],
                                                         IN2 := #space,
                                                         IN3 := #stringBox[#pString]);
                       END_IF;
                   END_REGION

                   REGION "TEST STRING NOT TOO LONG"
                       IF LEN(#lengthTest) <= #maxLength THEN
                           #_lineBox[#pLineBox] := #lengthTest;
                       END_IF;
                   END_REGION

                   REGION "TEST STRING TOO LONG"
                       IF LEN(#lengthTest) > #maxLength THEN
                           #_lineBox[#pLineBox] := "Trim"(#_lineBox[#pLineBox]);
                           #_lineBox[#pLineBox] := "Trim"(#_lineBox[#pLineBox]);
                           #pLineBox := #pLineBox + 1;
                           #_lineBox[#pLineBox] := #stringBox[#pString];
                       END_IF;
                   END_REGION

               END_IF;
           END_REGION

       END_FOR;
   END_REGION

   REGION "RETURN"
       #lineBox := #_lineBox;
   END_REGION
END_FUNCTION

